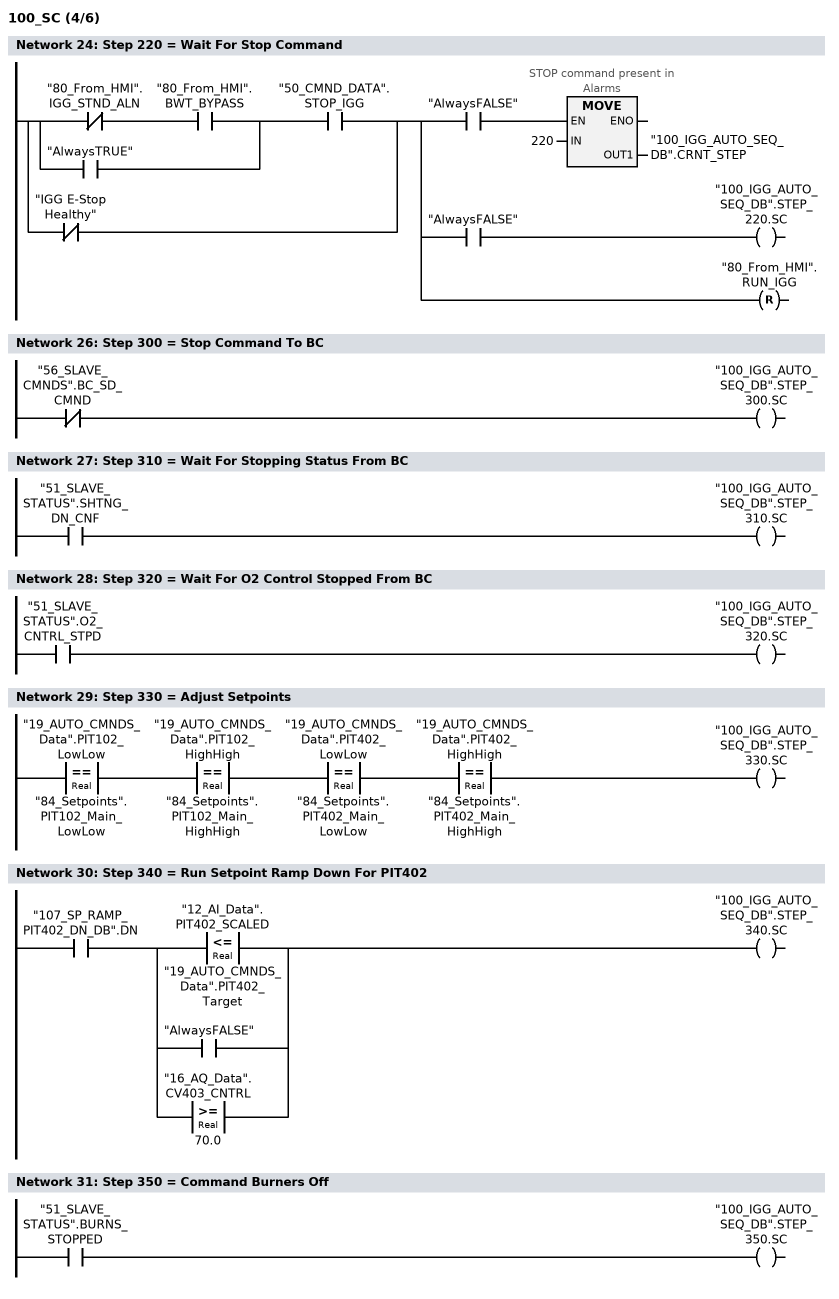
   RUNG wire#powerrail
      I_Contact( "80_From_HMI".IGG_STND_ALN )
      Contact( "80_From_HMI".BWT_BYPASS )
      wire#w1
      Contact( "50_CMND_DATA".STOP_IGG )
      wire#w2
      Contact( "AlwaysFALSE" )
      Move(in := 220, out1 => "100_IGG_AUTO_SEQ_DB".CRNT_STEP)   // STOP command present in Alarms
   END_RUNG
   RUNG wire#powerrail
      Contact( "AlwaysTRUE" )
   END_RUNG wire#w1
   RUNG wire#powerrail
      I_Contact( "IGG E-Stop Healthy" )
   END_RUNG wire#w2
   RUNG wire#w2
      Contact( "AlwaysFALSE" )
      Coil( "100_IGG_AUTO_SEQ_DB".STEP_220.SC )
   END_RUNG
   RUNG wire#w2
      R_Coil( "80_From_HMI".RUN_IGG )
   END_RUNG
   // the same network as SCL:
   #_w1 := (((NOT "80_From_HMI".IGG_STND_ALN AND "80_From_HMI".BWT_BYPASS) OR "AlwaysTRUE") AND "50_CMND_DATA".STOP_IGG) OR NOT "IGG E-Stop Healthy";
   IF #_w1 AND "AlwaysFALSE" THEN
       "100_IGG_AUTO_SEQ_DB".CRNT_STEP := 220;   // STOP command present in Alarms
   END_IF;
   "100_IGG_AUTO_SEQ_DB".STEP_220.SC := #_w1 AND "AlwaysFALSE";
   IF #_w1 THEN "80_From_HMI".RUN_IGG := FALSE; END_IF;
END_REGION

REGION Network 26: Step 300 = Stop Command To BC
   RUNG wire#powerrail
      I_Contact( "56_SLAVE_CMNDS".BC_SD_CMND )
      Coil( "100_IGG_AUTO_SEQ_DB".STEP_300.SC )
   END_RUNG
   // the same network as SCL:
   "100_IGG_AUTO_SEQ_DB".STEP_300.SC := NOT "56_SLAVE_CMNDS".BC_SD_CMND;
END_REGION

REGION Network 27: Step 310 = Wait For Stopping Status From BC
   RUNG wire#powerrail
      Contact( "51_SLAVE_STATUS".SHTNG_DN_CNF )
      Coil( "100_IGG_AUTO_SEQ_DB".STEP_310.SC )
   END_RUNG
   // the same network as SCL:
   "100_IGG_AUTO_SEQ_DB".STEP_310.SC := "51_SLAVE_STATUS".SHTNG_DN_CNF;
END_REGION

REGION Network 28: Step 320 = Wait For O2 Control Stopped From BC
   RUNG wire#powerrail
      Contact( "51_SLAVE_STATUS".O2_CNTRL_STPD )
      Coil( "100_IGG_AUTO_SEQ_DB".STEP_320.SC )
   END_RUNG
   // the same network as SCL:
   "100_IGG_AUTO_SEQ_DB".STEP_320.SC := "51_SLAVE_STATUS".O2_CNTRL_STPD;
END_REGION

REGION Network 29: Step 330 = Adjust Setpoints
   RUNG wire#powerrail
      { S7_Templates := "SrcType := Real" } EQ_Contact(in1 := "19_AUTO_CMNDS_Data".PIT102_LowLow, in2 := "84_Setpoints".PIT102_Main_LowLow)
      { S7_Templates := "SrcType := Real" } EQ_Contact(in1 := "19_AUTO_CMNDS_Data".PIT102_HighHigh, in2 := "84_Setpoints".PIT102_Main_HighHigh)
      { S7_Templates := "SrcType := Real" } EQ_Contact(in1 := "19_AUTO_CMNDS_Data".PIT402_LowLow, in2 := "84_Setpoints".PIT402_Main_LowLow)
      { S7_Templates := "SrcType := Real" } EQ_Contact(in1 := "19_AUTO_CMNDS_Data".PIT402_HighHigh, in2 := "84_Setpoints".PIT402_Main_HighHigh)
      Coil( "100_IGG_AUTO_SEQ_DB".STEP_330.SC )
   END_RUNG
   // the same network as SCL:
   "100_IGG_AUTO_SEQ_DB".STEP_330.SC := ("19_AUTO_CMNDS_Data".PIT102_LowLow = "84_Setpoints".PIT102_Main_LowLow) AND ("19_AUTO_CMNDS_Data".PIT102_HighHigh = "84_Setpoints".PIT102_Main_HighHigh) AND ("19_AUTO_CMNDS_Data".PIT402_LowLow = "84_Setpoints".PIT402_Main_LowLow) AND ("19_AUTO_CMNDS_Data".PIT402_HighHigh = "84_Setpoints".PIT402_Main_HighHigh);
END_REGION

REGION Network 30: Step 340 = Run Setpoint Ramp Down For PIT402
   RUNG wire#powerrail
      Contact( "107_SP_RAMP_PIT402_DN_DB".DN )
      wire#w1
      { S7_Templates := "SrcType := Real" } LE_Contact(in1 := "12_AI_Data".PIT402_SCALED, in2 := "19_AUTO_CMNDS_Data".PIT402_Target)
      wire#w2
      Coil( "100_IGG_AUTO_SEQ_DB".STEP_340.SC )
   END_RUNG
   RUNG wire#w1
      Contact( "AlwaysFALSE" )
   END_RUNG wire#w2
   RUNG wire#w1
      { S7_Templates := "SrcType := Real" } GE_Contact(in1 := "16_AQ_Data".CV403_CNTRL, in2 := 70.0)
   END_RUNG wire#w2
   // the same network as SCL:
   "100_IGG_AUTO_SEQ_DB".STEP_340.SC := "107_SP_RAMP_PIT402_DN_DB".DN AND (("12_AI_Data".PIT402_SCALED <= "19_AUTO_CMNDS_Data".PIT402_Target) OR "AlwaysFALSE" OR ("16_AQ_Data".CV403_CNTRL >= 70.0));
END_REGION

REGION Network 31: Step 350 = Command Burners Off
   RUNG wire#powerrail
      Contact( "51_SLAVE_STATUS".BURNS_STOPPED )
      Coil( "100_IGG_AUTO_SEQ_DB".STEP_350.SC )
   END_RUNG
   // the same network as SCL:
   "100_IGG_AUTO_SEQ_DB".STEP_350.SC := "51_SLAVE_STATUS".BURNS_STOPPED;
END_REGION

REGION Network 32: Step 360 = CV403 To 100% (Fully Open)
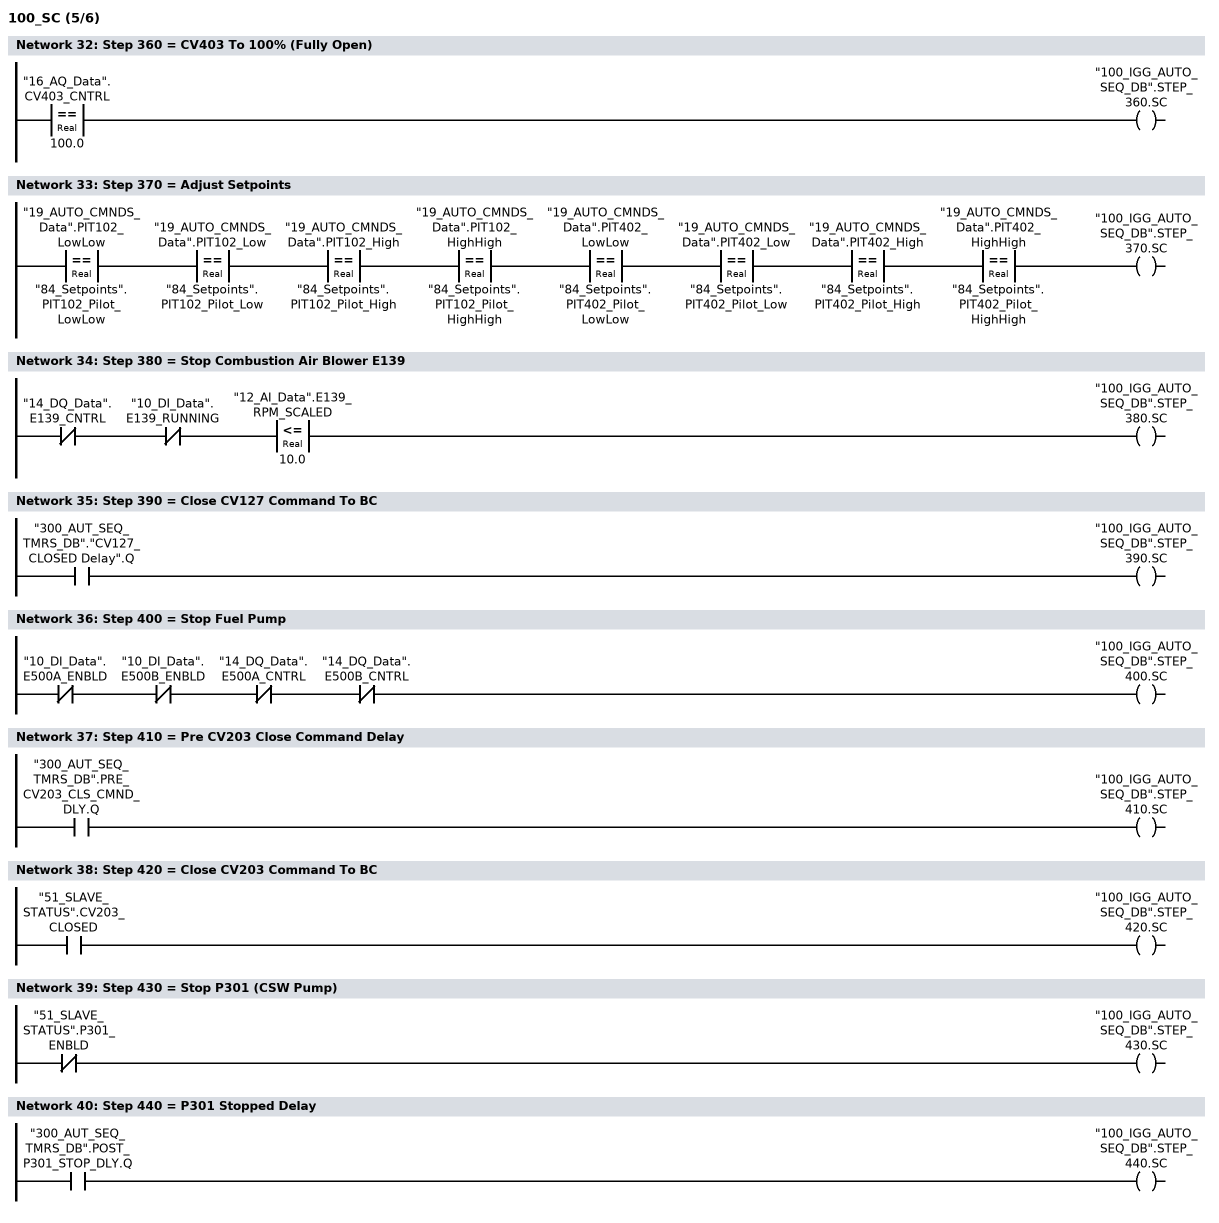
   RUNG wire#powerrail
      { S7_Templates := "SrcType := Real" } EQ_Contact(in1 := "16_AQ_Data".CV403_CNTRL, in2 := 100.0)
      Coil( "100_IGG_AUTO_SEQ_DB".STEP_360.SC )
   END_RUNG
   // the same network as SCL:
   "100_IGG_AUTO_SEQ_DB".STEP_360.SC := "16_AQ_Data".CV403_CNTRL = 100.0;
END_REGION

REGION Network 33: Step 370 = Adjust Setpoints
   RUNG wire#powerrail
      { S7_Templates := "SrcType := Real" } EQ_Contact(in1 := "19_AUTO_CMNDS_Data".PIT102_LowLow, in2 := "84_Setpoints".PIT102_Pilot_LowLow)
      { S7_Templates := "SrcType := Real" } EQ_Contact(in1 := "19_AUTO_CMNDS_Data".PIT102_Low, in2 := "84_Setpoints".PIT102_Pilot_Low)
      { S7_Templates := "SrcType := Real" } EQ_Contact(in1 := "19_AUTO_CMNDS_Data".PIT102_High, in2 := "84_Setpoints".PIT102_Pilot_High)
      { S7_Templates := "SrcType := Real" } EQ_Contact(in1 := "19_AUTO_CMNDS_Data".PIT102_HighHigh, in2 := "84_Setpoints".PIT102_Pilot_HighHigh)
      { S7_Templates := "SrcType := Real" } EQ_Contact(in1 := "19_AUTO_CMNDS_Data".PIT402_LowLow, in2 := "84_Setpoints".PIT402_Pilot_LowLow)
      { S7_Templates := "SrcType := Real" } EQ_Contact(in1 := "19_AUTO_CMNDS_Data".PIT402_Low, in2 := "84_Setpoints".PIT402_Pilot_Low)
      { S7_Templates := "SrcType := Real" } EQ_Contact(in1 := "19_AUTO_CMNDS_Data".PIT402_High, in2 := "84_Setpoints".PIT402_Pilot_High)
      { S7_Templates := "SrcType := Real" } EQ_Contact(in1 := "19_AUTO_CMNDS_Data".PIT402_HighHigh, in2 := "84_Setpoints".PIT402_Pilot_HighHigh)
      Coil( "100_IGG_AUTO_SEQ_DB".STEP_370.SC )
   END_RUNG
   // the same network as SCL:
   "100_IGG_AUTO_SEQ_DB".STEP_370.SC := ("19_AUTO_CMNDS_Data".PIT102_LowLow = "84_Setpoints".PIT102_Pilot_LowLow) AND ("19_AUTO_CMNDS_Data".PIT102_Low = "84_Setpoints".PIT102_Pilot_Low) AND ("19_AUTO_CMNDS_Data".PIT102_High = "84_Setpoints".PIT102_Pilot_High) AND ("19_AUTO_CMNDS_Data".PIT102_HighHigh = "84_Setpoints".PIT102_Pilot_HighHigh) AND ("19_AUTO_CMNDS_Data".PIT402_LowLow = "84_Setpoints".PIT402_Pilot_LowLow) AND ("19_AUTO_CMNDS_Data".PIT402_Low = "84_Setpoints".PIT402_Pilot_Low) AND ("19_AUTO_CMNDS_Data".PIT402_High = "84_Setpoints".PIT402_Pilot_High) AND ("19_AUTO_CMNDS_Data".PIT402_HighHigh = "84_Setpoints".PIT402_Pilot_HighHigh);
END_REGION

REGION Network 34: Step 380 = Stop Combustion Air Blower E139
   RUNG wire#powerrail
      I_Contact( "14_DQ_Data".E139_CNTRL )
      I_Contact( "10_DI_Data".E139_RUNNING )
      { S7_Templates := "SrcType := Real" } LE_Contact(in1 := "12_AI_Data".E139_RPM_SCALED, in2 := 10.0)
      Coil( "100_IGG_AUTO_SEQ_DB".STEP_380.SC )
   END_RUNG
   // the same network as SCL:
   "100_IGG_AUTO_SEQ_DB".STEP_380.SC := NOT "14_DQ_Data".E139_CNTRL AND NOT "10_DI_Data".E139_RUNNING AND ("12_AI_Data".E139_RPM_SCALED <= 10.0);
END_REGION

REGION Network 35: Step 390 = Close CV127 Command To BC
   RUNG wire#powerrail
      Contact( "300_AUT_SEQ_TMRS_DB"."CV127_CLOSED Delay".Q )
      Coil( "100_IGG_AUTO_SEQ_DB".STEP_390.SC )
   END_RUNG
   // the same network as SCL:
   "100_IGG_AUTO_SEQ_DB".STEP_390.SC := "300_AUT_SEQ_TMRS_DB"."CV127_CLOSED Delay".Q;
END_REGION

REGION Network 36: Step 400 = Stop Fuel Pump
   RUNG wire#powerrail
      I_Contact( "10_DI_Data".E500A_ENBLD )
      I_Contact( "10_DI_Data".E500B_ENBLD )
      I_Contact( "14_DQ_Data".E500A_CNTRL )
      I_Contact( "14_DQ_Data".E500B_CNTRL )
      Coil( "100_IGG_AUTO_SEQ_DB".STEP_400.SC )
   END_RUNG
   // the same network as SCL:
   "100_IGG_AUTO_SEQ_DB".STEP_400.SC := NOT "10_DI_Data".E500A_ENBLD AND NOT "10_DI_Data".E500B_ENBLD AND NOT "14_DQ_Data".E500A_CNTRL AND NOT "14_DQ_Data".E500B_CNTRL;
END_REGION

REGION Network 37: Step 410 = Pre CV203 Close Command Delay
   RUNG wire#powerrail
      Contact( "300_AUT_SEQ_TMRS_DB".PRE_CV203_CLS_CMND_DLY.Q )
      Coil( "100_IGG_AUTO_SEQ_DB".STEP_410.SC )
   END_RUNG
   // the same network as SCL:
   "100_IGG_AUTO_SEQ_DB".STEP_410.SC := "300_AUT_SEQ_TMRS_DB".PRE_CV203_CLS_CMND_DLY.Q;
END_REGION

REGION Network 38: Step 420 = Close CV203 Command To BC
   RUNG wire#powerrail
      Contact( "51_SLAVE_STATUS".CV203_CLOSED )
      Coil( "100_IGG_AUTO_SEQ_DB".STEP_420.SC )
   END_RUNG
   // the same network as SCL:
   "100_IGG_AUTO_SEQ_DB".STEP_420.SC := "51_SLAVE_STATUS".CV203_CLOSED;
END_REGION

REGION Network 39: Step 430 = Stop P301 (CSW Pump)
   RUNG wire#powerrail
      I_Contact( "51_SLAVE_STATUS".P301_ENBLD )
      Coil( "100_IGG_AUTO_SEQ_DB".STEP_430.SC )
   END_RUNG
   // the same network as SCL:
   "100_IGG_AUTO_SEQ_DB".STEP_430.SC := NOT "51_SLAVE_STATUS".P301_ENBLD;
END_REGION

REGION Network 40: Step 440 = P301 Stopped Delay
   RUNG wire#powerrail
      Contact( "300_AUT_SEQ_TMRS_DB".POST_P301_STOP_DLY.Q )
      Coil( "100_IGG_AUTO_SEQ_DB".STEP_440.SC )
   END_RUNG
   // the same network as SCL:
   "100_IGG_AUTO_SEQ_DB".STEP_440.SC := "300_AUT_SEQ_TMRS_DB".POST_P301_STOP_DLY.Q;
END_REGION

REGION Network 41: Step 450 = Cooling Water inlet Valves To Initial Position CV311 = Closed & CV312 = Open
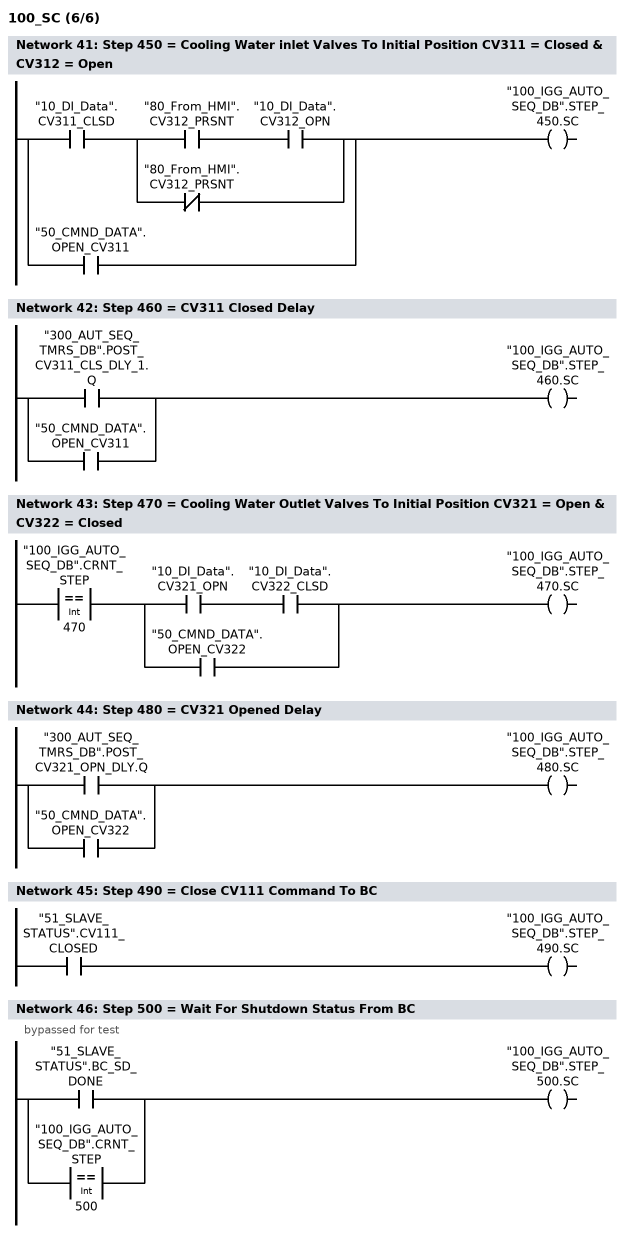
   RUNG wire#powerrail
      Contact( "10_DI_Data".CV311_CLSD )
      wire#w1
      Contact( "80_From_HMI".CV312_PRSNT )
      Contact( "10_DI_Data".CV312_OPN )
      wire#w2
      Coil( "100_IGG_AUTO_SEQ_DB".STEP_450.SC )
   END_RUNG
   RUNG wire#w1
      I_Contact( "80_From_HMI".CV312_PRSNT )
   END_RUNG wire#w2
   RUNG wire#powerrail
      Contact( "50_CMND_DATA".OPEN_CV311 )
   END_RUNG wire#w2
   // the same network as SCL:
   "100_IGG_AUTO_SEQ_DB".STEP_450.SC := ("10_DI_Data".CV311_CLSD AND (("80_From_HMI".CV312_PRSNT AND "10_DI_Data".CV312_OPN) OR NOT "80_From_HMI".CV312_PRSNT)) OR "50_CMND_DATA".OPEN_CV311;
END_REGION

REGION Network 42: Step 460 = CV311 Closed Delay
   RUNG wire#powerrail
      Contact( "300_AUT_SEQ_TMRS_DB".POST_CV311_CLS_DLY_1.Q )
      wire#w1
      Coil( "100_IGG_AUTO_SEQ_DB".STEP_460.SC )
   END_RUNG
   RUNG wire#powerrail
      Contact( "50_CMND_DATA".OPEN_CV311 )
   END_RUNG wire#w1
   // the same network as SCL:
   "100_IGG_AUTO_SEQ_DB".STEP_460.SC := "300_AUT_SEQ_TMRS_DB".POST_CV311_CLS_DLY_1.Q OR "50_CMND_DATA".OPEN_CV311;
END_REGION

REGION Network 43: Step 470 = Cooling Water Outlet Valves To Initial Position CV321 = Open & CV322 = Closed
   RUNG wire#powerrail
      { S7_Templates := "SrcType := Int" } EQ_Contact(in1 := "100_IGG_AUTO_SEQ_DB".CRNT_STEP, in2 := 470)
      wire#w1
      Contact( "10_DI_Data".CV321_OPN )
      Contact( "10_DI_Data".CV322_CLSD )
      wire#w2
      Coil( "100_IGG_AUTO_SEQ_DB".STEP_470.SC )
   END_RUNG
   RUNG wire#w1
      Contact( "50_CMND_DATA".OPEN_CV322 )
   END_RUNG wire#w2
   // the same network as SCL:
   "100_IGG_AUTO_SEQ_DB".STEP_470.SC := ("100_IGG_AUTO_SEQ_DB".CRNT_STEP = 470) AND (("10_DI_Data".CV321_OPN AND "10_DI_Data".CV322_CLSD) OR "50_CMND_DATA".OPEN_CV322);
END_REGION

REGION Network 44: Step 480 = CV321 Opened Delay
   RUNG wire#powerrail
      Contact( "300_AUT_SEQ_TMRS_DB".POST_CV321_OPN_DLY.Q )
      wire#w1
      Coil( "100_IGG_AUTO_SEQ_DB".STEP_480.SC )
   END_RUNG
   RUNG wire#powerrail
      Contact( "50_CMND_DATA".OPEN_CV322 )
   END_RUNG wire#w1
   // the same network as SCL:
   "100_IGG_AUTO_SEQ_DB".STEP_480.SC := "300_AUT_SEQ_TMRS_DB".POST_CV321_OPN_DLY.Q OR "50_CMND_DATA".OPEN_CV322;
END_REGION

REGION Network 45: Step 490 = Close CV111 Command To BC
   RUNG wire#powerrail
      Contact( "51_SLAVE_STATUS".CV111_CLOSED )
      Coil( "100_IGG_AUTO_SEQ_DB".STEP_490.SC )
   END_RUNG
   // the same network as SCL:
   "100_IGG_AUTO_SEQ_DB".STEP_490.SC := "51_SLAVE_STATUS".CV111_CLOSED;
END_REGION

REGION Network 46: Step 500 = Wait For Shutdown Status From BC
   // bypassed for test
   RUNG wire#powerrail
      Contact( "51_SLAVE_STATUS".BC_SD_DONE )
      wire#w1
      Coil( "100_IGG_AUTO_SEQ_DB".STEP_500.SC )
   END_RUNG
   RUNG wire#powerrail
      { S7_Templates := "SrcType := Int" } EQ_Contact(in1 := "100_IGG_AUTO_SEQ_DB".CRNT_STEP, in2 := 500)
   END_RUNG wire#w1
   // the same network as SCL:
   "100_IGG_AUTO_SEQ_DB".STEP_500.SC := "51_SLAVE_STATUS".BC_SD_DONE OR ("100_IGG_AUTO_SEQ_DB".CRNT_STEP = 500);
END_REGION
END_FUNCTION

FUNCTION "101_SP_CNFG" : Void   // FC101, LAD
TITLE = Setpoint Configuration
{ S7_Optimized_Access := 'TRUE' }
AUTHOR : JRS
VERSION : 0.1
// For configuring setpoints during automatic operation
   VAR_TEMP   // added for the SCL form of the ladder/FBD networks
      _w1 : Bool;
   END_VAR
BEGIN

REGION Network 1: PIT402 Setpoints
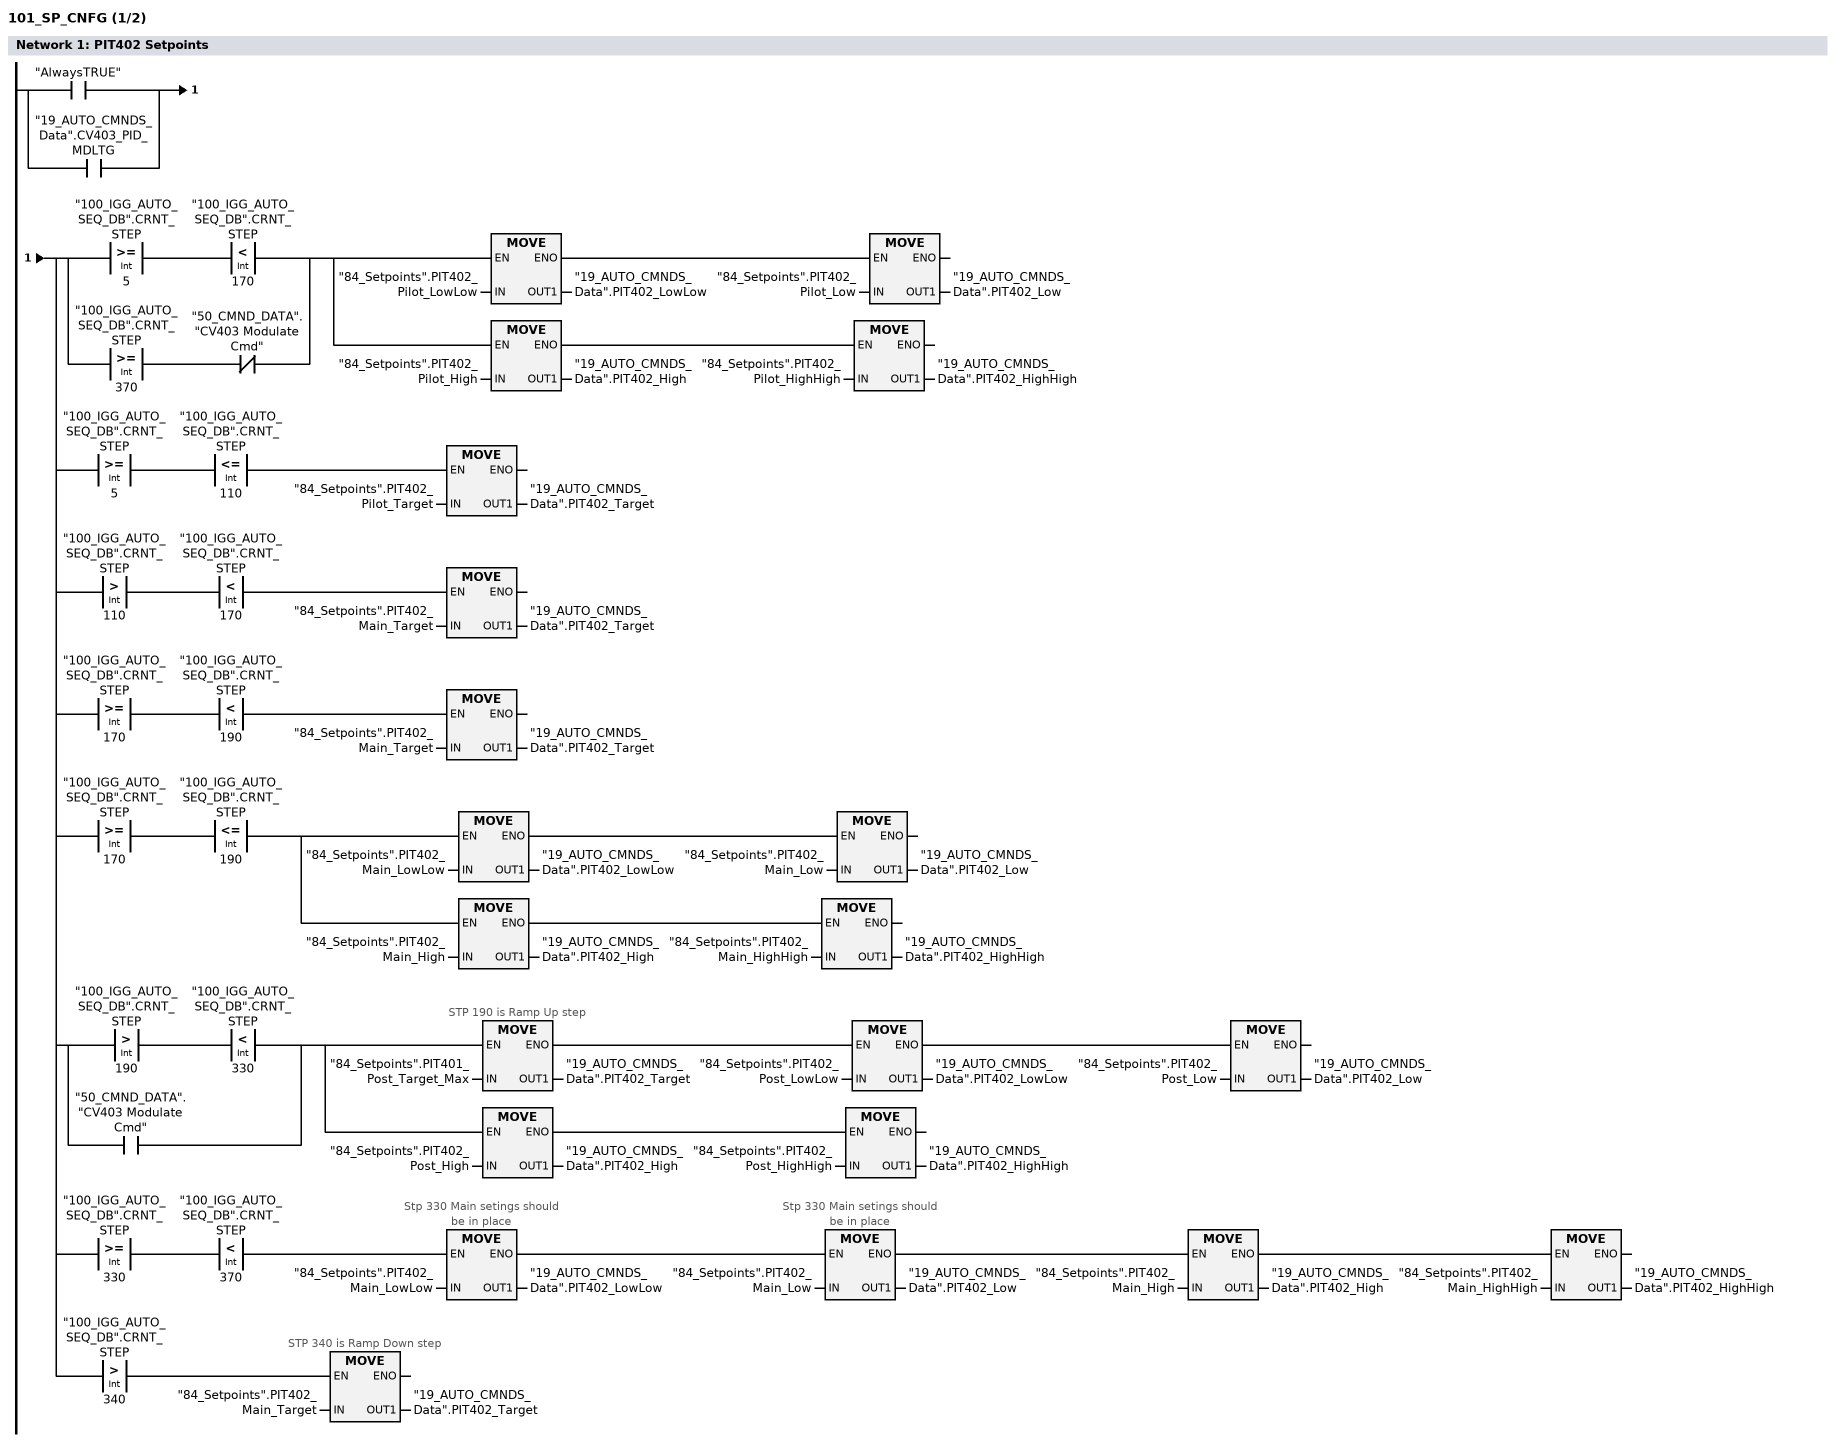
   RUNG wire#powerrail
      Contact( "AlwaysTRUE" )
      wire#w1
      { S7_Templates := "SrcType := Int" } GE_Contact(in1 := "100_IGG_AUTO_SEQ_DB".CRNT_STEP, in2 := 5)
      { S7_Templates := "SrcType := Int" } LT_Contact(in1 := "100_IGG_AUTO_SEQ_DB".CRNT_STEP, in2 := 170)
      wire#w2
      Move(in := "84_Setpoints".PIT402_Pilot_LowLow, out1 => "19_AUTO_CMNDS_Data".PIT402_LowLow)
      Move(in := "84_Setpoints".PIT402_Pilot_Low, out1 => "19_AUTO_CMNDS_Data".PIT402_Low)
   END_RUNG
   RUNG wire#powerrail
      Contact( "19_AUTO_CMNDS_Data".CV403_PID_MDLTG )
   END_RUNG wire#w1
   RUNG wire#w1
      { S7_Templates := "SrcType := Int" } GE_Contact(in1 := "100_IGG_AUTO_SEQ_DB".CRNT_STEP, in2 := 370)
      I_Contact( "50_CMND_DATA"."CV403 Modulate Cmd" )
   END_RUNG wire#w2
   RUNG wire#w2
      Move(in := "84_Setpoints".PIT402_Pilot_High, out1 => "19_AUTO_CMNDS_Data".PIT402_High)
      Move(in := "84_Setpoints".PIT402_Pilot_HighHigh, out1 => "19_AUTO_CMNDS_Data".PIT402_HighHigh)
   END_RUNG
   RUNG wire#w1
      { S7_Templates := "SrcType := Int" } GE_Contact(in1 := "100_IGG_AUTO_SEQ_DB".CRNT_STEP, in2 := 5)
      { S7_Templates := "SrcType := Int" } LE_Contact(in1 := "100_IGG_AUTO_SEQ_DB".CRNT_STEP, in2 := 110)
      Move(in := "84_Setpoints".PIT402_Pilot_Target, out1 => "19_AUTO_CMNDS_Data".PIT402_Target)
   END_RUNG
   RUNG wire#w1
      { S7_Templates := "SrcType := Int" } GT_Contact(in1 := "100_IGG_AUTO_SEQ_DB".CRNT_STEP, in2 := 110)
      { S7_Templates := "SrcType := Int" } LT_Contact(in1 := "100_IGG_AUTO_SEQ_DB".CRNT_STEP, in2 := 170)
      Move(in := "84_Setpoints".PIT402_Main_Target, out1 => "19_AUTO_CMNDS_Data".PIT402_Target)
   END_RUNG
   RUNG wire#w1
      { S7_Templates := "SrcType := Int" } GE_Contact(in1 := "100_IGG_AUTO_SEQ_DB".CRNT_STEP, in2 := 170)
      { S7_Templates := "SrcType := Int" } LT_Contact(in1 := "100_IGG_AUTO_SEQ_DB".CRNT_STEP, in2 := 190)
      Move(in := "84_Setpoints".PIT402_Main_Target, out1 => "19_AUTO_CMNDS_Data".PIT402_Target)
   END_RUNG
   RUNG wire#w1
      { S7_Templates := "SrcType := Int" } GE_Contact(in1 := "100_IGG_AUTO_SEQ_DB".CRNT_STEP, in2 := 170)
      { S7_Templates := "SrcType := Int" } LE_Contact(in1 := "100_IGG_AUTO_SEQ_DB".CRNT_STEP, in2 := 190)
      wire#w3
      Move(in := "84_Setpoints".PIT402_Main_LowLow, out1 => "19_AUTO_CMNDS_Data".PIT402_LowLow)
      Move(in := "84_Setpoints".PIT402_Main_Low, out1 => "19_AUTO_CMNDS_Data".PIT402_Low)
   END_RUNG
   RUNG wire#w3
      Move(in := "84_Setpoints".PIT402_Main_High, out1 => "19_AUTO_CMNDS_Data".PIT402_High)
      Move(in := "84_Setpoints".PIT402_Main_HighHigh, out1 => "19_AUTO_CMNDS_Data".PIT402_HighHigh)
   END_RUNG
   RUNG wire#w1
      { S7_Templates := "SrcType := Int" } GT_Contact(in1 := "100_IGG_AUTO_SEQ_DB".CRNT_STEP, in2 := 190)
      { S7_Templates := "SrcType := Int" } LT_Contact(in1 := "100_IGG_AUTO_SEQ_DB".CRNT_STEP, in2 := 330)
      wire#w4
      Move(in := "84_Setpoints".PIT401_Post_Target_Max, out1 => "19_AUTO_CMNDS_Data".PIT402_Target)   // STP 190 is Ramp Up step
      Move(in := "84_Setpoints".PIT402_Post_LowLow, out1 => "19_AUTO_CMNDS_Data".PIT402_LowLow)
      Move(in := "84_Setpoints".PIT402_Post_Low, out1 => "19_AUTO_CMNDS_Data".PIT402_Low)
   END_RUNG
   RUNG wire#w1
      Contact( "50_CMND_DATA"."CV403 Modulate Cmd" )
   END_RUNG wire#w4
   RUNG wire#w4
      Move(in := "84_Setpoints".PIT402_Post_High, out1 => "19_AUTO_CMNDS_Data".PIT402_High)
      Move(in := "84_Setpoints".PIT402_Post_HighHigh, out1 => "19_AUTO_CMNDS_Data".PIT402_HighHigh)
   END_RUNG
   RUNG wire#w1
      { S7_Templates := "SrcType := Int" } GE_Contact(in1 := "100_IGG_AUTO_SEQ_DB".CRNT_STEP, in2 := 330)
      { S7_Templates := "SrcType := Int" } LT_Contact(in1 := "100_IGG_AUTO_SEQ_DB".CRNT_STEP, in2 := 370)
      Move(in := "84_Setpoints".PIT402_Main_LowLow, out1 => "19_AUTO_CMNDS_Data".PIT402_LowLow)   // Stp 330 Main setings should be in place
      Move(in := "84_Setpoints".PIT402_Main_Low, out1 => "19_AUTO_CMNDS_Data".PIT402_Low)   // Stp 330 Main setings should be in place
      Move(in := "84_Setpoints".PIT402_Main_High, out1 => "19_AUTO_CMNDS_Data".PIT402_High)
      Move(in := "84_Setpoints".PIT402_Main_HighHigh, out1 => "19_AUTO_CMNDS_Data".PIT402_HighHigh)
   END_RUNG
   RUNG wire#w1
      { S7_Templates := "SrcType := Int" } GT_Contact(in1 := "100_IGG_AUTO_SEQ_DB".CRNT_STEP, in2 := 340)
      Move(in := "84_Setpoints".PIT402_Main_Target, out1 => "19_AUTO_CMNDS_Data".PIT402_Target)   // STP 340 is Ramp Down step
   END_RUNG
   // the same network as SCL:
   #_w1 := "AlwaysTRUE" OR "19_AUTO_CMNDS_Data".CV403_PID_MDLTG;
   IF #_w1 AND ((("100_IGG_AUTO_SEQ_DB".CRNT_STEP >= 5) AND ("100_IGG_AUTO_SEQ_DB".CRNT_STEP < 170)) OR (("100_IGG_AUTO_SEQ_DB".CRNT_STEP >= 370) AND NOT "50_CMND_DATA"."CV403 Modulate Cmd")) THEN
       "19_AUTO_CMNDS_Data".PIT402_LowLow := "84_Setpoints".PIT402_Pilot_LowLow;
       "19_AUTO_CMNDS_Data".PIT402_Low := "84_Setpoints".PIT402_Pilot_Low;
       "19_AUTO_CMNDS_Data".PIT402_High := "84_Setpoints".PIT402_Pilot_High;
       "19_AUTO_CMNDS_Data".PIT402_HighHigh := "84_Setpoints".PIT402_Pilot_HighHigh;
   END_IF;
   IF #_w1 AND ("100_IGG_AUTO_SEQ_DB".CRNT_STEP >= 5) AND ("100_IGG_AUTO_SEQ_DB".CRNT_STEP <= 110) THEN
       "19_AUTO_CMNDS_Data".PIT402_Target := "84_Setpoints".PIT402_Pilot_Target;
   END_IF;
   IF #_w1 AND ("100_IGG_AUTO_SEQ_DB".CRNT_STEP > 110) AND ("100_IGG_AUTO_SEQ_DB".CRNT_STEP < 170) THEN
       "19_AUTO_CMNDS_Data".PIT402_Target := "84_Setpoints".PIT402_Main_Target;
   END_IF;
   IF #_w1 AND ("100_IGG_AUTO_SEQ_DB".CRNT_STEP >= 170) AND ("100_IGG_AUTO_SEQ_DB".CRNT_STEP < 190) THEN
       "19_AUTO_CMNDS_Data".PIT402_Target := "84_Setpoints".PIT402_Main_Target;
   END_IF;
   IF #_w1 AND ("100_IGG_AUTO_SEQ_DB".CRNT_STEP >= 170) AND ("100_IGG_AUTO_SEQ_DB".CRNT_STEP <= 190) THEN
       "19_AUTO_CMNDS_Data".PIT402_LowLow := "84_Setpoints".PIT402_Main_LowLow;
       "19_AUTO_CMNDS_Data".PIT402_Low := "84_Setpoints".PIT402_Main_Low;
       "19_AUTO_CMNDS_Data".PIT402_High := "84_Setpoints".PIT402_Main_High;
       "19_AUTO_CMNDS_Data".PIT402_HighHigh := "84_Setpoints".PIT402_Main_HighHigh;
   END_IF;
   IF #_w1 AND ((("100_IGG_AUTO_SEQ_DB".CRNT_STEP > 190) AND ("100_IGG_AUTO_SEQ_DB".CRNT_STEP < 330)) OR "50_CMND_DATA"."CV403 Modulate Cmd") THEN
       "19_AUTO_CMNDS_Data".PIT402_Target := "84_Setpoints".PIT401_Post_Target_Max;   // STP 190 is Ramp Up step
       "19_AUTO_CMNDS_Data".PIT402_LowLow := "84_Setpoints".PIT402_Post_LowLow;
       "19_AUTO_CMNDS_Data".PIT402_Low := "84_Setpoints".PIT402_Post_Low;
       "19_AUTO_CMNDS_Data".PIT402_High := "84_Setpoints".PIT402_Post_High;
       "19_AUTO_CMNDS_Data".PIT402_HighHigh := "84_Setpoints".PIT402_Post_HighHigh;
   END_IF;
   IF #_w1 AND ("100_IGG_AUTO_SEQ_DB".CRNT_STEP >= 330) AND ("100_IGG_AUTO_SEQ_DB".CRNT_STEP < 370) THEN
       "19_AUTO_CMNDS_Data".PIT402_LowLow := "84_Setpoints".PIT402_Main_LowLow;   // Stp 330 Main setings should be in place
       "19_AUTO_CMNDS_Data".PIT402_Low := "84_Setpoints".PIT402_Main_Low;   // Stp 330 Main setings should be in place
       "19_AUTO_CMNDS_Data".PIT402_High := "84_Setpoints".PIT402_Main_High;
       "19_AUTO_CMNDS_Data".PIT402_HighHigh := "84_Setpoints".PIT402_Main_HighHigh;
   END_IF;
   IF #_w1 AND ("100_IGG_AUTO_SEQ_DB".CRNT_STEP > 340) THEN
       "19_AUTO_CMNDS_Data".PIT402_Target := "84_Setpoints".PIT402_Main_Target;   // STP 340 is Ramp Down step
   END_IF;
END_REGION

REGION Network 2: PIT102 Setpoints
   // Changed from 130 to 5 for test  changed to 180 from 190